(* Logix 5000 project; controller MV vendor 1 type 14 code 217 rev 31.11; software revision 31.00; part 53 of 53 *)
(* tags used below, declared in another part *)
   Alarm_Reset : BOOL;
   Analog_Fault_No : DINT;
   Analog_Simulation_Enabled : BOOL;
   CWD : CHECKWORD_FLAGS;
   Default_Check_Time : DINT;
   Dummy : BOOL;
   Item_Faults_Are_Latched : BOOL;
   Item_Simulation_Flag : BOOL;
   ItoF_raw_input : INT;
   MV_B17 : INT[255];   // VES_ACTIVE Vessel active flags
   MV_bit_data_file_address : INT;
   mv_bit_file_bit_offset : INT;
   mv_bit_file_word_offset : INT;
   MV_bit_offset : INT;
   MV_bit_value_to_set : INT;
   MV_BM01_AV01 : PlantItem;   // BM01_AV01
   MV_BM01_AV01_ALARM : ALARM_DIGITAL;
   MV_BM01_AV01_C : ALIAS FOR Remote_IO:8:I.Data.6;
   MV_BM01_AV01_CIP : BOOL;
   MV_BM01_AV01_DR : ALIAS FOR Remote_IO:9:O.Data.3;
   MV_BM01_AV01_MV20 : BOOL;
   MV_BM01_AV01_MV21 : BOOL;
   MV_BM01_AV01_mv22 : BOOL;
   MV_BM01_AV01_O : ALIAS FOR Remote_IO:8:I.Data.7;
   MV_DAL01_AV01 : PlantItem;   // DAL01_AV01
   MV_DAL01_AV01_ALARM : ALARM_DIGITAL;
   MV_DAL01_AV01_C : ALIAS FOR Remote_IO:8:I.Data.8;
   MV_DAL01_AV01_DR : ALIAS FOR Remote_IO:9:O.Data.4;
   MV_DAL01_AV01_MV20 : BOOL;
   MV_DAL01_AV01_MV21 : BOOL;
   MV_DAL01_AV01_mv22 : BOOL;
   MV_DAL01_AV01_O : ALIAS FOR Remote_IO:8:I.Data.9;
   MV_data_file_address : INT;
   MV_Data_To_TF : DINT[30];
   MV_MV20_AV01 : PlantItem;   // MV20_AV01
   MV_MV20_AV01_ALARM : ALARM_DIGITAL;
   MV_MV20_AV01_C : ALIAS FOR Remote_IO:8:I.Data.0;
   MV_MV20_AV01_DR : ALIAS FOR Remote_IO:9:O.Data.0;
   MV_MV20_AV01_O : ALIAS FOR Remote_IO:8:I.Data.1;
   MV_MV21_AV01 : PlantItem;   // MV21_AV01
   MV_MV21_AV01_ALARM : ALARM_DIGITAL;
   MV_MV21_AV01_C : ALIAS FOR Remote_IO:8:I.Data.2;
   MV_MV21_AV01_DR : ALIAS FOR Remote_IO:9:O.Data.1;
   MV_MV21_AV01_O : ALIAS FOR Remote_IO:8:I.Data.3;
   MV_MV22_AV01 : PlantItem;   // MV22_AV01
   MV_MV22_AV01_ALARM : ALARM_DIGITAL;
   MV_MV22_AV01_C : ALIAS FOR Remote_IO:8:I.Data.4;
   MV_MV22_AV01_DR : ALIAS FOR Remote_IO:9:O.Data.2;
   MV_MV22_AV01_O : ALIAS FOR Remote_IO:8:I.Data.5;
   One_Second_One_Scan : ALIAS FOR One_Second_1_scan;
   overrange_RIO_analog_value : REAL;
   rack_simulation_flag : BOOL;
   Scada_Pump_Fault_No : DINT;
   Scada_Pump_H_Fault_No : DINT;
   Scada_Pump_T_Fault_No : DINT;
   Scada_Valve_Fault_No : DINT;
   scale_analog_int : DINT;
   scale_analog_result : REAL;
   scale_eu_max : REAL;
   scale_eu_min : REAL;
   scale_raw_input : REAL;
   scale_raw_max : REAL;
   scale_raw_min : REAL;
   scale_routine_active : BOOL;
   scale_temp : REAL;
   template_analog_input : PlantItem;
   template_analog_input_RawInput : REAL;
   template_analog_output : PlantItem;
   template_analog_output_RawOutput : REAL;
   template_input : PlantItem;
   template_input_RawInput : ALIAS FOR template_boolean;
   template_output : PlantItem;
   template_output_RawOutput : ALIAS FOR template_boolean;   // P04CHILLRUN Chiller Run Signal
   template_pump : PlantItem;
   template_pump_D : ALIAS FOR template_boolean;   // auto start vacuum pump 1
   template_pump_ISOL : ALIAS FOR template_boolean;
   template_pump_R : ALIAS FOR template_boolean;   // vacuum pump 1 running
   template_valve : PlantItem;
   template_valve_C : ALIAS FOR template_boolean;   // skim manifold to ycv2 drain valve closed
   template_valve_DR : ALIAS FOR template_boolean;   // drive open skim manifold to ycv2 drain valve
   template_valve_O : ALIAS FOR template_boolean;   // skim manifold to ycv2 drain valve opened
   underrange_RIO_analog_value : REAL;
(* MV_Common, continued *)

ROUTINE MV_SetBitFile_Value   (* ladder *)
   // Sets the Value of a bit within a bit file, Can use complete bit offset across words
   0: SBR(MV_bit_value_to_set,MV_bit_data_file_address,MV_bit_offset)OTE(Dummy);
   1: DIV(MV_data_file_address,16,mv_bit_file_word_offset)MOD(MV_data_file_address,16,mv_bit_file_bit_offset);
   // Bit File 17
   2: EQU(MV_bit_data_file_address,17)[EQU(MV_bit_value_to_set,1) OTL(MV_B17[mv_bit_file_word_offset].[mv_bit_file_bit_offset]) ,EQU(MV_bit_value_to_set,0) OTU(MV_B17[mv_bit_file_word_offset].[mv_bit_file_bit_offset]) ];
   3: RET();
END_ROUTINE

ROUTINE MV_Valves   (* ladder *)
   0: [NEQ(MV_MV20_AV01.DriveBits,0) OTE(MV_MV20_AV01.CW.[CWD.AUTODRV]) ,[XIC(MV_MV20_AV01.CW.[CWD.AUTODRV]) XIO(MV_MV20_AV01.CW.[CWD.MANUAL]) ,XIC(MV_MV20_AV01.CW.[CWD.MANDRV]) XIC(MV_MV20_AV01.CW.[CWD.MANUAL]) ] OTE(MV_MV20_AV01.CW.[CWD.OUTPUT]) ,XIC(MV_MV20_AV01.CW.[CWD.OUTPUT]) OTE(MV_MV20_AV01_DR) ,XIC(S:FS) [OTU(MV_MV20_AV01.CW.[CWD.MANUAL]) ,LEQ(MV_MV20_AV01.CheckTime,0) MOV(Default_Check_Time,MV_MV20_AV01.CheckTime) ] ,[[XIC(MV_MV20_AV01_O) XIO(Item_Simulation_Flag) ,XIC(Item_Simulation_Flag) XIC(MV_MV20_AV01.CW.[CWD.OUTPUT]) XIO(MV_MV20_AV01.CW.[CWD.SIMFAIL]) ] OTE(MV_MV20_AV01.CW.[CWD.OPENFB]) ,[XIC(MV_MV20_AV01_C) XIO(Item_Simulation_Flag) ,XIC(Item_Simulation_Flag) XIO(MV_MV20_AV01.CW.[CWD.OUTPUT]) XIO(MV_MV20_AV01.CW.[CWD.SIMFAIL]) ] OTE(MV_MV20_AV01.CW.[CWD.CLOSEDFB]) ] ,[XIC(MV_MV20_AV01.CW.[CWD.OUTPUT]) XIO(MV_MV20_AV01.CW.[CWD.PREVSCAN]) ,XIO(MV_MV20_AV01.CW.[CWD.OUTPUT]) XIC(MV_MV20_AV01.CW.[CWD.PREVSCAN]) ] CLR(MV_MV20_AV01.CheckTimer) ,XIC(One_Second_One_Scan) LES(MV_MV20_AV01.CheckTimer,MV_MV20_AV01.CheckTime) ADD(MV_MV20_AV01.CheckTimer,1,MV_MV20_AV01.CheckTimer) ,XIO(MV_MV20_AV01.CW.[CWD.FAULT]) OTU(MV_MV20_AV01.CW.[CWD.FAULTLOGGED]) ,[GEQ(MV_MV20_AV01.CheckTimer,MV_MV20_AV01.CheckTime) [XIC(MV_MV20_AV01.CW.[CWD.OUTPUT]) [XIO(MV_MV20_AV01.CW.[CWD.OPENFB]) ,XIC(MV_MV20_AV01.CW.[CWD.CLOSEDFB]) ] ,XIO(MV_MV20_AV01.CW.[CWD.OUTPUT]) [XIC(MV_MV20_AV01.CW.[CWD.OPENFB]) ,XIO(MV_MV20_AV01.CW.[CWD.CLOSEDFB]) ] ] ,XIC(MV_MV20_AV01.CW.[CWD.FAULT]) XIC(Item_Faults_Are_Latched) ,XIC(MV_MV20_AV01.CW.[CWD.HIGHLIGHT]) ] XIO(MV_MV20_AV01.CW.[CWD.CHECKOFF]) XIO(Alarm_Reset) [OTE(MV_MV20_AV01.CW.[CWD.FAULT]) ,ALMD(MV_MV20_AV01_ALARM,0,0,0,0) ] ,XIC(MV_MV20_AV01.CW.[CWD.OUTPUT]) OTE(MV_MV20_AV01.CW.[CWD.PREVSCAN]) ];
   1: [NEQ(MV_MV21_AV01.DriveBits,0) OTE(MV_MV21_AV01.CW.[CWD.AUTODRV]) ,[XIC(MV_MV21_AV01.CW.[CWD.AUTODRV]) XIO(MV_MV21_AV01.CW.[CWD.MANUAL]) ,XIC(MV_MV21_AV01.CW.[CWD.MANDRV]) XIC(MV_MV21_AV01.CW.[CWD.MANUAL]) ] OTE(MV_MV21_AV01.CW.[CWD.OUTPUT]) ,XIC(MV_MV21_AV01.CW.[CWD.OUTPUT]) OTE(MV_MV21_AV01_DR) ,XIC(S:FS) [OTU(MV_MV21_AV01.CW.[CWD.MANUAL]) ,LEQ(MV_MV21_AV01.CheckTime,0) MOV(Default_Check_Time,MV_MV21_AV01.CheckTime) ] ,[[XIC(MV_MV21_AV01_O) XIO(Item_Simulation_Flag) ,XIC(Item_Simulation_Flag) XIC(MV_MV21_AV01.CW.[CWD.OUTPUT]) XIO(MV_MV21_AV01.CW.[CWD.SIMFAIL]) ] OTE(MV_MV21_AV01.CW.[CWD.OPENFB]) ,[XIC(MV_MV21_AV01_C) XIO(Item_Simulation_Flag) ,XIC(Item_Simulation_Flag) XIO(MV_MV21_AV01.CW.[CWD.OUTPUT]) XIO(MV_MV21_AV01.CW.[CWD.SIMFAIL]) ] OTE(MV_MV21_AV01.CW.[CWD.CLOSEDFB]) ] ,[XIC(MV_MV21_AV01.CW.[CWD.OUTPUT]) XIO(MV_MV21_AV01.CW.[CWD.PREVSCAN]) ,XIO(MV_MV21_AV01.CW.[CWD.OUTPUT]) XIC(MV_MV21_AV01.CW.[CWD.PREVSCAN]) ] CLR(MV_MV21_AV01.CheckTimer) ,XIC(One_Second_One_Scan) LES(MV_MV21_AV01.CheckTimer,MV_MV21_AV01.CheckTime) ADD(MV_MV21_AV01.CheckTimer,1,MV_MV21_AV01.CheckTimer) ,XIO(MV_MV21_AV01.CW.[CWD.FAULT]) OTU(MV_MV21_AV01.CW.[CWD.FAULTLOGGED]) ,[GEQ(MV_MV21_AV01.CheckTimer,MV_MV21_AV01.CheckTime) [XIC(MV_MV21_AV01.CW.[CWD.OUTPUT]) [XIO(MV_MV21_AV01.CW.[CWD.OPENFB]) ,XIC(MV_MV21_AV01.CW.[CWD.CLOSEDFB]) ] ,XIO(MV_MV21_AV01.CW.[CWD.OUTPUT]) [XIC(MV_MV21_AV01.CW.[CWD.OPENFB]) ,XIO(MV_MV21_AV01.CW.[CWD.CLOSEDFB]) ] ] ,XIC(MV_MV21_AV01.CW.[CWD.FAULT]) XIC(Item_Faults_Are_Latched) ,XIC(MV_MV21_AV01.CW.[CWD.HIGHLIGHT]) ] XIO(MV_MV21_AV01.CW.[CWD.CHECKOFF]) XIO(Alarm_Reset) [OTE(MV_MV21_AV01.CW.[CWD.FAULT]) ,ALMD(MV_MV21_AV01_ALARM,0,0,0,0) ] ,XIC(MV_MV21_AV01.CW.[CWD.OUTPUT]) OTE(MV_MV21_AV01.CW.[CWD.PREVSCAN]) ];
   2: [NEQ(MV_MV22_AV01.DriveBits,0) OTE(MV_MV22_AV01.CW.[CWD.AUTODRV]) ,[XIC(MV_MV22_AV01.CW.[CWD.AUTODRV]) XIO(MV_MV22_AV01.CW.[CWD.MANUAL]) ,XIC(MV_MV22_AV01.CW.[CWD.MANDRV]) XIC(MV_MV22_AV01.CW.[CWD.MANUAL]) ] OTE(MV_MV22_AV01.CW.[CWD.OUTPUT]) ,XIC(MV_MV22_AV01.CW.[CWD.OUTPUT]) OTE(MV_MV22_AV01_DR) ,XIC(S:FS) [OTU(MV_MV22_AV01.CW.[CWD.MANUAL]) ,LEQ(MV_MV22_AV01.CheckTime,0) MOV(Default_Check_Time,MV_MV22_AV01.CheckTime) ] ,[[XIC(MV_MV22_AV01_O) XIO(Item_Simulation_Flag) ,XIC(Item_Simulation_Flag) XIC(MV_MV22_AV01.CW.[CWD.OUTPUT]) XIO(MV_MV22_AV01.CW.[CWD.SIMFAIL]) ] OTE(MV_MV22_AV01.CW.[CWD.OPENFB]) ,[XIC(MV_MV22_AV01_C) XIO(Item_Simulation_Flag) ,XIC(Item_Simulation_Flag) XIO(MV_MV22_AV01.CW.[CWD.OUTPUT]) XIO(MV_MV22_AV01.CW.[CWD.SIMFAIL]) ] OTE(MV_MV22_AV01.CW.[CWD.CLOSEDFB]) ] ,[XIC(MV_MV22_AV01.CW.[CWD.OUTPUT]) XIO(MV_MV22_AV01.CW.[CWD.PREVSCAN]) ,XIO(MV_MV22_AV01.CW.[CWD.OUTPUT]) XIC(MV_MV22_AV01.CW.[CWD.PREVSCAN]) ] CLR(MV_MV22_AV01.CheckTimer) ,XIC(One_Second_One_Scan) LES(MV_MV22_AV01.CheckTimer,MV_MV22_AV01.CheckTime) ADD(MV_MV22_AV01.CheckTimer,1,MV_MV22_AV01.CheckTimer) ,XIO(MV_MV22_AV01.CW.[CWD.FAULT]) OTU(MV_MV22_AV01.CW.[CWD.FAULTLOGGED]) ,[GEQ(MV_MV22_AV01.CheckTimer,MV_MV22_AV01.CheckTime) [XIC(MV_MV22_AV01.CW.[CWD.OUTPUT]) [XIO(MV_MV22_AV01.CW.[CWD.OPENFB]) ,XIC(MV_MV22_AV01.CW.[CWD.CLOSEDFB]) ] ,XIO(MV_MV22_AV01.CW.[CWD.OUTPUT]) [XIC(MV_MV22_AV01.CW.[CWD.OPENFB]) ,XIO(MV_MV22_AV01.CW.[CWD.CLOSEDFB]) ] ] ,XIC(MV_MV22_AV01.CW.[CWD.FAULT]) XIC(Item_Faults_Are_Latched) ,XIC(MV_MV22_AV01.CW.[CWD.HIGHLIGHT]) ] XIO(MV_MV22_AV01.CW.[CWD.CHECKOFF]) XIO(Alarm_Reset) [OTE(MV_MV22_AV01.CW.[CWD.FAULT]) ,ALMD(MV_MV22_AV01_ALARM,0,0,0,0) ] ,XIC(MV_MV22_AV01.CW.[CWD.OUTPUT]) OTE(MV_MV22_AV01.CW.[CWD.PREVSCAN]) ];
   3: [XIC(MV_BM01_AV01_MV20) ,XIC(MV_BM01_AV01_MV21) ,XIC(MV_BM01_AV01_mv22) ,XIC(MV_BM01_AV01_CIP) ]OTE(MV_BM01_AV01.DriveBits.0);
   4: [NEQ(MV_BM01_AV01.DriveBits,0) OTE(MV_BM01_AV01.CW.[CWD.AUTODRV]) ,[XIC(MV_BM01_AV01.CW.[CWD.AUTODRV]) XIO(MV_BM01_AV01.CW.[CWD.MANUAL]) ,XIC(MV_BM01_AV01.CW.[CWD.MANDRV]) XIC(MV_BM01_AV01.CW.[CWD.MANUAL]) ] OTE(MV_BM01_AV01.CW.[CWD.OUTPUT]) ,XIC(MV_BM01_AV01.CW.[CWD.OUTPUT]) OTE(MV_BM01_AV01_DR) ,XIC(S:FS) [OTU(MV_BM01_AV01.CW.[CWD.MANUAL]) ,LEQ(MV_BM01_AV01.CheckTime,0) MOV(Default_Check_Time,MV_BM01_AV01.CheckTime) ] ,[[XIC(MV_BM01_AV01_O) XIO(Item_Simulation_Flag) ,XIC(Item_Simulation_Flag) XIC(MV_BM01_AV01.CW.[CWD.OUTPUT]) XIO(MV_BM01_AV01.CW.[CWD.SIMFAIL]) ] [OTE(MV_BM01_AV01.CW.[CWD.OPENFB]) ,OTE(MV_Data_To_TF[2].0) ] ,[XIC(MV_BM01_AV01_C) XIO(Item_Simulation_Flag) ,XIC(Item_Simulation_Flag) XIO(MV_BM01_AV01.CW.[CWD.OUTPUT]) XIO(MV_BM01_AV01.CW.[CWD.SIMFAIL]) ] OTE(MV_BM01_AV01.CW.[CWD.CLOSEDFB]) ] ,[XIC(MV_BM01_AV01.CW.[CWD.OUTPUT]) XIO(MV_BM01_AV01.CW.[CWD.PREVSCAN]) ,XIO(MV_BM01_AV01.CW.[CWD.OUTPUT]) XIC(MV_BM01_AV01.CW.[CWD.PREVSCAN]) ] CLR(MV_BM01_AV01.CheckTimer) ,XIC(One_Second_One_Scan) LES(MV_BM01_AV01.CheckTimer,MV_BM01_AV01.CheckTime) ADD(MV_BM01_AV01.CheckTimer,1,MV_BM01_AV01.CheckTimer) ,XIO(MV_BM01_AV01.CW.[CWD.FAULT]) OTU(MV_BM01_AV01.CW.[CWD.FAULTLOGGED]) ,[GEQ(MV_BM01_AV01.CheckTimer,MV_BM01_AV01.CheckTime) [XIC(MV_BM01_AV01.CW.[CWD.OUTPUT]) [XIO(MV_BM01_AV01.CW.[CWD.OPENFB]) ,XIC(MV_BM01_AV01.CW.[CWD.CLOSEDFB]) ] ,XIO(MV_BM01_AV01.CW.[CWD.OUTPUT]) [XIC(MV_BM01_AV01.CW.[CWD.OPENFB]) ,XIO(MV_BM01_AV01.CW.[CWD.CLOSEDFB]) ] ] ,XIC(MV_BM01_AV01.CW.[CWD.FAULT]) XIC(Item_Faults_Are_Latched) ,XIC(MV_BM01_AV01.CW.[CWD.HIGHLIGHT]) ] XIO(MV_BM01_AV01.CW.[CWD.CHECKOFF]) XIO(Alarm_Reset) [OTE(MV_BM01_AV01.CW.[CWD.FAULT]) ,ALMD(MV_BM01_AV01_ALARM,0,0,0,0) ] ,XIC(MV_BM01_AV01.CW.[CWD.OUTPUT]) OTE(MV_BM01_AV01.CW.[CWD.PREVSCAN]) ];
   5: [XIC(MV_DAL01_AV01_MV20) ,XIC(MV_DAL01_AV01_MV21) ,XIC(MV_DAL01_AV01_mv22) ]OTE(MV_DAL01_AV01.DriveBits.0);
   6: [NEQ(MV_DAL01_AV01.DriveBits,0) OTE(MV_DAL01_AV01.CW.[CWD.AUTODRV]) ,[XIC(MV_DAL01_AV01.CW.[CWD.AUTODRV]) XIO(MV_DAL01_AV01.CW.[CWD.MANUAL]) ,XIC(MV_DAL01_AV01.CW.[CWD.MANDRV]) XIC(MV_DAL01_AV01.CW.[CWD.MANUAL]) ] OTE(MV_DAL01_AV01.CW.[CWD.OUTPUT]) ,XIC(MV_DAL01_AV01.CW.[CWD.OUTPUT]) OTE(MV_DAL01_AV01_DR) ,XIC(S:FS) [OTU(MV_DAL01_AV01.CW.[CWD.MANUAL]) ,LEQ(MV_DAL01_AV01.CheckTime,0) MOV(Default_Check_Time,MV_DAL01_AV01.CheckTime) ] ,[[XIC(MV_DAL01_AV01_O) XIO(Item_Simulation_Flag) ,XIC(Item_Simulation_Flag) XIC(MV_DAL01_AV01.CW.[CWD.OUTPUT]) XIO(MV_DAL01_AV01.CW.[CWD.SIMFAIL]) ] [OTE(MV_DAL01_AV01.CW.[CWD.OPENFB]) ,OTE(MV_Data_To_TF[0].0) ] ,[XIC(MV_DAL01_AV01_C) XIO(Item_Simulation_Flag) ,XIC(Item_Simulation_Flag) XIO(MV_DAL01_AV01.CW.[CWD.OUTPUT]) XIO(MV_DAL01_AV01.CW.[CWD.SIMFAIL]) ] OTE(MV_DAL01_AV01.CW.[CWD.CLOSEDFB]) ] ,[XIC(MV_DAL01_AV01.CW.[CWD.OUTPUT]) XIO(MV_DAL01_AV01.CW.[CWD.PREVSCAN]) ,XIO(MV_DAL01_AV01.CW.[CWD.OUTPUT]) XIC(MV_DAL01_AV01.CW.[CWD.PREVSCAN]) ] CLR(MV_DAL01_AV01.CheckTimer) ,XIC(One_Second_One_Scan) LES(MV_DAL01_AV01.CheckTimer,MV_DAL01_AV01.CheckTime) ADD(MV_DAL01_AV01.CheckTimer,1,MV_DAL01_AV01.CheckTimer) ,XIO(MV_DAL01_AV01.CW.[CWD.FAULT]) OTU(MV_DAL01_AV01.CW.[CWD.FAULTLOGGED]) ,[GEQ(MV_DAL01_AV01.CheckTimer,MV_DAL01_AV01.CheckTime) [XIC(MV_DAL01_AV01.CW.[CWD.OUTPUT]) [XIO(MV_DAL01_AV01.CW.[CWD.OPENFB]) ,XIC(MV_DAL01_AV01.CW.[CWD.CLOSEDFB]) ] ,XIO(MV_DAL01_AV01.CW.[CWD.OUTPUT]) [XIC(MV_DAL01_AV01.CW.[CWD.OPENFB]) ,XIO(MV_DAL01_AV01.CW.[CWD.CLOSEDFB]) ] ] ,XIC(MV_DAL01_AV01.CW.[CWD.FAULT]) XIC(Item_Faults_Are_Latched) ,XIC(MV_DAL01_AV01.CW.[CWD.HIGHLIGHT]) ] XIO(MV_DAL01_AV01.CW.[CWD.CHECKOFF]) XIO(Alarm_Reset) [OTE(MV_DAL01_AV01.CW.[CWD.FAULT]) ,ALMD(MV_DAL01_AV01_ALARM,0,0,0,0) ] ,XIC(MV_DAL01_AV01.CW.[CWD.OUTPUT]) OTE(MV_DAL01_AV01.CW.[CWD.PREVSCAN]) ];
END_ROUTINE
END_PROGRAM

PROGRAM Templates   (* main routine Normal_Input_Template *)

ROUTINE Analog_Scale_FtoI   (* ladder *)
   0: SBR(scale_raw_input,scale_raw_min,scale_raw_max,scale_eu_min,scale_eu_max)OTE(scale_routine_active);
   1: CPT(scale_temp,(scale_eu_max-scale_eu_min)/(scale_raw_max-scale_raw_min));
   2: CPT(scale_analog_result,(scale_raw_input-scale_raw_min)*scale_temp+scale_eu_min);
   3: ADD(scale_analog_result,0.0,scale_analog_int);
   4: RET(scale_analog_int);
END_ROUTINE

ROUTINE Analog_Scale_ItoF   (* ladder *)
   0: SBR(ItoF_raw_input,scale_raw_min,scale_raw_max,scale_eu_min,scale_eu_max)OTE(scale_routine_active);
   1: ADD(ItoF_raw_input,0.0,scale_raw_input);
   2: CPT(scale_temp,(scale_eu_max-scale_eu_min)/(scale_raw_max-scale_raw_min));
   3: CPT(scale_analog_result,(scale_raw_input-scale_raw_min)*scale_temp+scale_eu_min);
   4: RET(scale_analog_result);
END_ROUTINE

ROUTINE Normal_Analogue_Input   (* ladder *)
   0: XIO(Analog_Simulation_Enabled)[XIO(template_analog_input.CW.[CWD.MANUAL]) JSR(Analog_Scale_ItoF,5,template_analog_input_RawInput,0.0,30840.0,0.0,6500.0,template_analog_input.Scaled) ,[LIM(underrange_RIO_analog_value,template_analog_input_RawInput,overrange_RIO_analog_value) ,XIC(template_analog_input.CW.[CWD.CHECKOFF]) ] CLR(template_analog_input.CheckTimer) ,XIC(S:FS) [OTU(template_analog_input.CW.[CWD.MANUAL]) ,LEQ(template_analog_input.CheckTime,0) MOV(Default_Check_Time,template_analog_input.CheckTime) ] ,XIC(One_Second_One_Scan) LES(template_analog_input.CheckTimer,template_analog_input.CheckTime) ADD(template_analog_input.CheckTimer,1,template_analog_input.CheckTimer) ,GEQ(template_analog_input.CheckTimer,template_analog_input.CheckTime) XIO(Alarm_Reset) OTE(template_analog_input.CW.[CWD.FAULT]) ,XIC(template_analog_input.CW.[CWD.FAULT]) EQU(Analog_Fault_No,0) XIO(template_analog_input.CW.[CWD.FAULTLOGGED]) [MOV(30001,Analog_Fault_No) ,OTL(template_analog_input.CW.[CWD.FAULTLOGGED]) ] ];
END_ROUTINE

ROUTINE Normal_Analogue_Output   (* ladder *)
   0: XIO(Analog_Simulation_Enabled)JSR(Analog_Scale_FtoI,5,template_analog_output.Scaled,0.0,100.0,0.0,30840.0,template_analog_output_RawOutput);
END_ROUTINE

ROUTINE Normal_Input_Template   (* ladder *)
   0: [XIC(S:FS) OTU(template_input.CW.[CWD.MANUAL]) ,[XIC(template_input_RawInput) XIO(template_input.CW.[CWD.MANUAL]) ,XIC(template_input.CW.[CWD.MANDRV]) XIC(template_input.CW.[CWD.MANUAL]) ] OTE(template_input.CW.[CWD.INPUTSTATUS]) ,XIC(One_Second_One_Scan) [XIC(template_input.CW.[CWD.INPUTSTATUS]) XIO(template_input.CW.[CWD.INPUTSTATUSDEBOUNCED]) ,XIO(template_input.CW.[CWD.INPUTSTATUS]) XIC(template_input.CW.[CWD.INPUTSTATUSDEBOUNCED]) ] ADD(1,template_input.DebounceTimer,template_input.DebounceTimer) ,[XIC(template_input.CW.[CWD.INPUTSTATUS]) XIC(template_input.CW.[CWD.INPUTSTATUSDEBOUNCED]) ,XIO(template_input.CW.[CWD.INPUTSTATUS]) XIO(template_input.CW.[CWD.INPUTSTATUSDEBOUNCED]) ] CLR(template_input.DebounceTimer) ,GEQ(template_input.DebounceTimer,template_input.DebounceTime) XIC(template_input.CW.[CWD.INPUTSTATUS]) [OTL(template_input.CW.[CWD.INPUTSTATUSDEBOUNCED]) ,CLR(template_input.DebounceTimer) ] ,GEQ(template_input.DebounceTimer,template_input.DebounceTime) XIO(template_input.CW.[CWD.INPUTSTATUS]) [OTU(template_input.CW.[CWD.INPUTSTATUSDEBOUNCED]) ,CLR(template_input.DebounceTimer) ] ];
END_ROUTINE

ROUTINE Normal_Output_Template   (* ladder *)
   0: [NEQ(template_output.DriveBits,0) OTE(template_output.CW.[CWD.AUTODRV]) ,XIC(S:FS) OTU(template_output.CW.[CWD.MANUAL]) ,[XIC(template_output.CW.[CWD.AUTODRV]) XIO(template_output.CW.[CWD.MANUAL]) ,XIC(template_output.CW.[CWD.MANDRV]) XIC(template_output.CW.[CWD.MANUAL]) ] OTE(template_output.CW.[CWD.OUTPUT]) ,XIC(template_output.CW.[CWD.OUTPUT]) OTE(template_output_RawOutput) ];
END_ROUTINE

ROUTINE Normal_Pump_Template_Isol   (* ladder *)
   0: [NEQ(template_pump.DriveBits,0) OTE(template_pump.CW.[CWD.AUTODRV]) ,[XIC(template_pump.CW.[CWD.AUTODRV]) XIO(template_pump.CW.[CWD.MANUAL]) ,XIC(template_pump.CW.[CWD.MANDRV]) XIC(template_pump.CW.[CWD.MANUAL]) ] OTE(template_pump.CW.[CWD.OUTPUT]) ,XIC(template_pump.CW.[CWD.OUTPUT]) OTE(template_pump_D) ,XIC(S:FS) [OTU(template_pump.CW.[CWD.MANUAL]) ,LEQ(template_pump.CheckTime,0) MOV(Default_Check_Time,template_pump.CheckTime) ] ,[[XIC(template_pump_R) XIO(Item_Simulation_Flag) ,XIC(Item_Simulation_Flag) [XIC(template_pump.CW.[CWD.AUTODRV]) XIO(template_pump.CW.[CWD.SIMFAIL]) ,XIO(template_pump.CW.[CWD.AUTODRV]) XIC(template_pump.CW.[CWD.SIMFAIL]) ] ] OTE(template_pump.CW.[CWD.RUNFB]) ,[XIC(rack_simulation_flag) ,XIC(template_pump.CW.[CWD.CHECKOFF]) ,XIC(template_pump_ISOL) ] OTE(template_pump.CW.[CWD.HEALTHYFB]) ] ,[XIC(template_pump.CW.[CWD.AUTODRV]) XIO(template_pump.CW.[CWD.PREVSCAN]) ,XIO(template_pump.CW.[CWD.AUTODRV]) XIC(template_pump.CW.[CWD.PREVSCAN]) ] CLR(template_pump.CheckTimer) ,XIC(One_Second_One_Scan) LES(template_pump.CheckTimer,template_pump.CheckTime) ADD(template_pump.CheckTimer,1,template_pump.CheckTimer) ,XIO(template_pump.CW.[CWD.FAULT]) OTU(template_pump.CW.[CWD.FAULTLOGGED]) ,[GEQ(template_pump.CheckTimer,template_pump.CheckTime) [XIC(template_pump.CW.[CWD.OUTPUT]) XIO(template_pump.CW.[CWD.RUNFB]) ,XIO(template_pump.CW.[CWD.OUTPUT]) XIC(template_pump.CW.[CWD.RUNFB]) ] ,XIO(template_pump.CW.[CWD.HEALTHYFB]) ,XIC(template_pump.CW.[CWD.FAULT]) ,XIC(template_pump.CW.[CWD.HIGHLIGHT]) ] XIO(template_pump.CW.[CWD.CHECKOFF]) XIO(Alarm_Reset) OTE(template_pump.CW.[CWD.FAULT]) ,XIC(template_pump.CW.[CWD.OUTPUT]) OTE(template_pump.CW.[CWD.PREVSCAN]) ,XIC(template_pump.CW.[CWD.FAULT]) EQU(Scada_Pump_Fault_No,0) XIO(template_pump.CW.[CWD.FAULTLOGGED]) [MOV(20001,Scada_Pump_Fault_No) ,OTL(template_pump.CW.[CWD.FAULTLOGGED]) ] ,XIO(template_pump.CW.[CWD.HEALTHYFB]) EQU(Scada_Pump_H_Fault_No,0) XIO(template_pump.CW.[CWD.HEALTHYFAULTLOGGED]) [MOV(20001,Scada_Pump_H_Fault_No) ,OTL(template_pump.CW.[CWD.HEALTHYFAULTLOGGED]) ] ,XIO(template_pump.CW.[CWD.NOTTRIPPEDFB]) EQU(Scada_Pump_H_Fault_No,0) XIO(template_pump.CW.[CWD.TRIPPEDFAULTLOGGED]) [MOV(20001,Scada_Pump_T_Fault_No) ,OTL(template_pump.CW.[CWD.TRIPPEDFAULTLOGGED]) ] ];
END_ROUTINE

ROUTINE Normal_Pump_Template_JustRun   (* ladder *)
   0: [NEQ(template_pump.DriveBits,0) OTE(template_pump.CW.[CWD.AUTODRV]) ,[XIC(template_pump.CW.[CWD.AUTODRV]) XIO(template_pump.CW.[CWD.MANUAL]) ,XIC(template_pump.CW.[CWD.MANDRV]) XIC(template_pump.CW.[CWD.MANUAL]) ] OTE(template_pump.CW.[CWD.OUTPUT]) ,XIC(template_pump.CW.[CWD.OUTPUT]) OTE(template_pump_D) ,XIC(S:FS) [OTU(template_pump.CW.[CWD.MANUAL]) ,LEQ(template_pump.CheckTime,0) MOV(Default_Check_Time,template_pump.CheckTime) ] ,[[XIC(template_pump_R) XIO(Item_Simulation_Flag) ,XIC(Item_Simulation_Flag) [XIC(template_pump.CW.[CWD.AUTODRV]) XIO(template_pump.CW.[CWD.SIMFAIL]) ,XIO(template_pump.CW.[CWD.AUTODRV]) XIC(template_pump.CW.[CWD.SIMFAIL]) ] ] OTE(template_pump.CW.[CWD.RUNFB]) ,[XIC(rack_simulation_flag) ,XIC(template_pump.CW.[CWD.CHECKOFF]) ,] OTE(template_pump.CW.[CWD.HEALTHYFB]) ] ,[XIC(template_pump.CW.[CWD.AUTODRV]) XIO(template_pump.CW.[CWD.PREVSCAN]) ,XIO(template_pump.CW.[CWD.AUTODRV]) XIC(template_pump.CW.[CWD.PREVSCAN]) ] CLR(template_pump.CheckTimer) ,XIC(One_Second_One_Scan) LES(template_pump.CheckTimer,template_pump.CheckTime) ADD(template_pump.CheckTimer,1,template_pump.CheckTimer) ,XIO(template_pump.CW.[CWD.FAULT]) OTU(template_pump.CW.[CWD.FAULTLOGGED]) ,[GEQ(template_pump.CheckTimer,template_pump.CheckTime) [XIC(template_pump.CW.[CWD.OUTPUT]) XIO(template_pump.CW.[CWD.RUNFB]) ,XIO(template_pump.CW.[CWD.OUTPUT]) XIC(template_pump.CW.[CWD.RUNFB]) ] ,XIO(template_pump.CW.[CWD.HEALTHYFB]) ,XIC(template_pump.CW.[CWD.FAULT]) ,XIC(template_pump.CW.[CWD.HIGHLIGHT]) ] XIO(template_pump.CW.[CWD.CHECKOFF]) XIO(Alarm_Reset) OTE(template_pump.CW.[CWD.FAULT]) ,XIC(template_pump.CW.[CWD.OUTPUT]) OTE(template_pump.CW.[CWD.PREVSCAN]) ,XIC(template_pump.CW.[CWD.FAULT]) EQU(Scada_Pump_Fault_No,0) XIO(template_pump.CW.[CWD.FAULTLOGGED]) [MOV(20001,Scada_Pump_Fault_No) ,OTL(template_pump.CW.[CWD.FAULTLOGGED]) ] ,XIO(template_pump.CW.[CWD.HEALTHYFB]) EQU(Scada_Pump_H_Fault_No,0) XIO(template_pump.CW.[CWD.HEALTHYFAULTLOGGED]) [MOV(20001,Scada_Pump_H_Fault_No) ,OTL(template_pump.CW.[CWD.HEALTHYFAULTLOGGED]) ] ,XIO(template_pump.CW.[CWD.NOTTRIPPEDFB]) EQU(Scada_Pump_H_Fault_No,0) XIO(template_pump.CW.[CWD.TRIPPEDFAULTLOGGED]) [MOV(20001,Scada_Pump_T_Fault_No) ,OTL(template_pump.CW.[CWD.TRIPPEDFAULTLOGGED]) ] ];
END_ROUTINE

ROUTINE Normal_Valve_Template   (* ladder *)
   0: [NEQ(template_valve.DriveBits,0) OTE(template_valve.CW.[CWD.AUTODRV]) ,[XIC(template_valve.CW.[CWD.AUTODRV]) XIO(template_valve.CW.[CWD.MANUAL]) ,XIC(template_valve.CW.[CWD.MANDRV]) XIC(template_valve.CW.[CWD.MANUAL]) ] OTE(template_valve.CW.[CWD.OUTPUT]) ,XIC(template_valve.CW.[CWD.OUTPUT]) OTE(template_valve_DR) ,XIC(S:FS) [OTU(template_valve.CW.[CWD.MANUAL]) ,LEQ(template_valve.CheckTime,0) MOV(Default_Check_Time,template_valve.CheckTime) ] ,[[XIC(template_valve_O) XIO(Item_Simulation_Flag) ,XIC(Item_Simulation_Flag) XIC(template_valve.CW.[CWD.AUTODRV]) XIO(template_valve.CW.[CWD.SIMFAIL]) ] OTE(template_valve.CW.[CWD.OPENFB]) ,[XIC(template_valve_C) XIO(Item_Simulation_Flag) ,XIC(Item_Simulation_Flag) XIO(template_valve.CW.[CWD.AUTODRV]) XIO(template_valve.CW.[CWD.SIMFAIL]) ] OTE(template_valve.CW.[CWD.CLOSEDFB]) ] ,[XIC(template_valve.CW.[CWD.AUTODRV]) XIO(template_valve.CW.[CWD.PREVSCAN]) ,XIO(template_valve.CW.[CWD.AUTODRV]) XIC(template_valve.CW.[CWD.PREVSCAN]) ] CLR(template_valve.CheckTimer) ,XIC(One_Second_One_Scan) LES(template_valve.CheckTimer,template_valve.CheckTime) ADD(template_valve.CheckTimer,1,template_valve.CheckTimer) ,XIO(template_valve.CW.[CWD.FAULT]) OTU(template_valve.CW.[CWD.FAULTLOGGED]) ,[GEQ(template_valve.CheckTimer,template_valve.CheckTime) [XIC(template_valve.CW.[CWD.OUTPUT]) [XIO(template_valve.CW.[CWD.OPENFB]) ,XIC(template_valve.CW.[CWD.CLOSEDFB]) ] ,XIO(template_valve.CW.[CWD.OUTPUT]) [XIC(template_valve.CW.[CWD.OPENFB]) ,XIO(template_valve.CW.[CWD.CLOSEDFB]) ] ] ,XIC(template_valve.CW.[CWD.FAULT]) ,XIC(template_valve.CW.[CWD.HIGHLIGHT]) ] XIO(template_valve.CW.[CWD.CHECKOFF]) XIO(Alarm_Reset) OTE(template_valve.CW.[CWD.FAULT]) ,XIC(template_valve.CW.[CWD.OUTPUT]) OTE(template_valve.CW.[CWD.PREVSCAN]) ,XIC(template_valve.CW.[CWD.FAULT]) EQU(Scada_Valve_Fault_No,0) XIO(template_valve.CW.[CWD.FAULTLOGGED]) [MOV(10001,Scada_Valve_Fault_No) ,OTL(template_valve.CW.[CWD.FAULTLOGGED]) ] ];
END_ROUTINE
END_PROGRAM
